      ProcessValue <- "84_Setpoints_PIT402_Main_Target"
   TextField "Text field_27" at 697,736 size 58x20; Text 'Opened'
   TextField "Text field_29" at 306,694 size 300x20; Text 'Air / Inert Gas Pressure Setpoint (Current)'
   AlarmView "Alarm view_1" at 0,777 size 1280x23
   TextField "Text field_6" at 531,373 size 64x18; Text 'Running'
   TextField "Text field_9" at 530,395 size 57x25; Text 'Running'
      Visibility <- "10_DI_Data_E139_RUNNING"
   IOField "I/O field_4" at 917,398 size 89x25; FormatPattern 999999; Unit h
      ProcessValue <- "82_To_HMI_CA Blower Total Run Hours"
   TextField "Text field_30" at 1011,400 size 123x20; Text 'Total Run Hours'
   IOField "I/O field_21" at 916,146 size 90x25; FormatPattern 999999; Unit  h
      ProcessValue <- "82_To_HMI_I&A Compressor Total Run Hours"
   TextField "Text field_31" at 1011,148 size 123x20; Text 'Total Run Hours'
   IOField "I/O field_22" at 935,109 size 40x25; FormatPattern 99; Unit d
      ProcessValue <- "82_To_HMI_P301 CSW Pump Run Days"
   IOField "I/O field_23" at 1068,362 size 40x25; FormatPattern 99; Unit s
      ProcessValue <- "82_To_HMI_CA Blower Run Seconds"

screen "Cooling System" 1280x800, template "Template"
   Group "Group_1" at 335,308 size 88x156; Picture "Graphic_148"
   Group "Group_2" at 298,412 size 194x121; Picture "Graphic_224"
   GraphicView "Graphic view_14" at 335,308 size 85x153; Picture "Graphic_148"
   GraphicView "Graphic view_9" at 298,414 size 189x119; Picture "Graphic_224"
   Group "Group_4" at 1043,404 size 88x156; Picture "Graphic_148"
   Group "Group_5" at 1006,508 size 194x121; Picture "Graphic_224"
   GraphicView "Graphic view_27" at 1043,404 size 85x153; Picture "Graphic_148"
   GraphicView "Graphic view_28" at 1006,511 size 189x119; Picture "Graphic_224"
   Rectangle "Rectangle_7" at 224,48 size 554x250
      Visibility <- "80_From_HMI_P301_PRSNT"
   GraphicView "Graphic view_13" at 501,485 size 115x33; Picture "Graphic_232"
   GraphicView "Graphic view_1" at 446,429 size 75x87; Picture "Graphic_238"
   GraphicView "Graphic view_34" at 489,470 size 52x87; Picture "Graphic_169"
   GraphicView "Graphic view_11" at 80,468 size 424x50; Picture "Graphic_232"
   Group "Group_3" at 298,308 size 194x225; Picture "Graphic_148"
   GraphicView "Graphic view_2" at 480,389 size 43x49; Picture "Graphic_231"
   GraphicView "Graphic view_23" at 832,606 size 29x189; Picture "Graphic_231"
   GraphicView "Graphic view_18" at 802,567 size 88x52; Picture "Graphic_240"
   GraphicView "Graphic view_7" at 175,602 size 43x189; Picture "Graphic_231"
   GraphicView "Graphic view_29" at 964,565 size 56x50; Picture "Graphic_232"
   GraphicView "Graphic view_16" at 1150,564 size 56x50; Picture "Graphic_232"
   GraphicView "Graphic view_10" at 175,547 size 43x16; Picture "Graphic_231"
   GraphicView "Graphic view_8" at 25,514 size 207x209; Picture "Graphic_230"
   Button "HmiScreenItemData_1" at 1,1 size 150x43; TextOn 'Back'; TextOff 'Main Index'
      on Release: ActivateScreen("02 Main Index", 0)
   Rectangle "Rectangle_8" at 237,87 size 528x35
      Visibility <- "80_From_HMI_P301_PRSNT"
   Button "Button_15" at 468,92 size 57x25; TextOn 'Enabled'; TextOff 'Disabled'
      Visibility <- "80_From_HMI_P301_PRSNT"
   Button "Button_16" at 622,92 size 64x25; TextOn 'Alarm'; TextOff 'Text'
      Visibility <- "80_From_HMI_P301_PRSNT"
   TextField "Text field_14" at 239,94 size 185x20; Text 'Cooling Sea Water Pump'
   Button "Button_1" at 545,92 size 57x25; TextOn 'Enabled'; TextOff 'Stopped'
      Visibility <- "80_From_HMI_P301_PRSNT"
   Rectangle "Rectangle_1" at 236,83 size 530x212
      Visibility <- "80_From_HMI_P301_PRSNT"
   TextField "Text field_1" at 387,56 size 235x26; Text 'Cooling System Control'
   TextField "Text field_32" at 468,92 size 57x25; Text 'Enabled'
      Visibility <- "10 DI_DATA_P301_ENBLD"
   TextField "Text field_2" at 543,92 size 59x25; Text 'Running'
      Visibility <- "10_DI_Data_CV311_OPN(1)"
   Button "Button_2" at 622,92 size 64x25; TextOn 'Alarm'; TextOff 'Tripped'
      Visibility <- "10 DI_DATA_P301_TRIPPED"
      Appearance <- "10 DI_DATA_P301_TRIPPED"
   TextField "Text field_72" at 2,524 size 121x38; Text 'Cooling Seawater Inlet'
   GraphicView "Graphic view_17" at 464,297 size 75x99; Picture "Graphic_229"
   GraphicView "Graphic view_4" at 801,333 size 43x255; Picture "Graphic_231"
   GraphicView "Graphic view_5" at 786,305 size 72x46; Picture "Graphic_234"
   GraphicView "Graphic view_6" at 25,472 size 56x43; Picture "Graphic_235"
   TextField "Text field_7" at 12,598 size 58x20; Text 'CV-312'
   TextField "Text field_33" at 352,317 size 54x22; Text 'Closed'
      Visibility <- "10_DI_Data_CV311_CLSD"
   TextField "Text field_3" at 352,317 size 54x22; Text 'Opened'
      Visibility <- "10_DI_Data_CV311_OPN"
   TextField "Text field_71" at 351,343 size 58x20; Text 'CV-311'
   GraphicView "Graphic view_3" at 159,470 size 75x87; Picture "Graphic_239"
   TextField "Text field_5" at 534,295 size 105x38; Text 'To Inert Gas Generator'
   TextField "Text field_69" at 13,624 size 54x22; Text 'Closed'
      Visibility <- "10_DI_Data_CV312_CLSD"
   TextField "Text field_6" at 853,250 size 125x55; Text 'Warm Water From Inert Gas Generator'
   GraphicView "Graphic view_31" at 248,441 size 24x34; Picture "Graphic_36"
   TextField "Text field_17" at 230,422 size 62x20; Text 'PIT-359'
   IOField "I/O field_6" at 226,403 size 68x18; FormatPattern 99.99; Unit  Bar
      ProcessValue <- "12_AI_Data_PIT359_SCALED"
   GraphicView "Graphic view_21" at 849,377 size 88x52; Picture "Graphic_241"
   GraphicView "Graphic view_22" at 848,417 size 43x157; Picture "Graphic_231"
   TextField "Text field_8" at 867,659 size 78x55; Text 'Drain To Oily Bilge Tank'
   GraphicView "Graphic view_25" at 896,422 size 43x134; Picture "Graphic_231"
   GraphicView "Graphic view_26" at 898,526 size 73x87; Picture "Graphic_242"
   Group "Group_6" at 1006,404 size 194x225; Picture "Graphic_148"
   TextField "Text field_12" at 1053,439 size 58x20; Text 'CV-322'
   TextField "Text field_13" at 1054,413 size 54x22; Text 'Closed'
      Visibility <- "10_DI_Data_CV322_CLSD"
   TextField "Text field_19" at 1054,413 size 54x22; Text 'Opened'
      Visibility <- "10_DI_Data_CV322_OPN"
   TextField "Text field_20" at 1190,615 size 88x38; Text 'To Overboard'
   GraphicView "Graphic view_24" at 697,598 size 181x170; Picture "Graphic_230"
   TextField "Text field_9" at 681,704 size 58x20; Text 'CV-321'
   TextField "Text field_11" at 682,678 size 54x22; Text 'Closed'
      Visibility <- "10_DI_Data_CV321_CLSD"
   GraphicView "Graphic view_15" at 244,714 size 40x61; Picture "Graphic_236"
   TextField "Text field_21" at 214,658 size 93x55; Text 'To Existing Flue Gas Scrubber'
   TextField "Text field_70" at 13,624 size 54x22; Text 'Opened'
      Visibility <- "10_DI_Data_CV312_OPN"
   TextField "Text field_10" at 682,678 size 54x22; Text 'Opened'
      Visibility <- "10_DI_Data_CV321_OPN"
   GraphicView "Graphic view_32" at 512,546 size 30x121; Picture "Graphic_147"
   TextField "Text field_4" at 600,529 size 79x55; Text 'Cooling Seawater To GCU'
   GraphicView "Graphic view_19" at 624,477 size 56x43; Picture "Graphic_235"
   GraphicView "Graphic view_33" at 508,659 size 40x61; Picture "Graphic_236"
   TextField "Text field_22" at 481,722 size 79x55; Text 'Cooling Seawater To PGC'
   GraphicView "Graphic view_12" at 891,714 size 40x61; Picture "Graphic_236"
   GraphicView "Graphic view_30" at 1206,568 size 56x43; Picture "Graphic_235"
   GraphicView "Graphic view_35" at 803,244 size 40x61; Picture "Graphic_236"
   Button "HmiScreenItemData_4" at 1129,1 size 150x43; TextOn 'I&A Compressor Ok'; TextOff 'Back'
      on Release: function_efd93a16()
   AlarmView "Alarm view_1" at 0,777 size 1280x23
   Button "HmiScreenItemData_11" at 345,230 size 69x51; TextOn 'RESET'; TextOff 'Reset'; Authorization "Operate"
      on Press: function_b14e0dd5("82_To_HMI_P301 CSW Pump Reset Hours", 0)
   IOField "I/O field_8" at 270,232 size 65x25; FormatPattern 99999; Unit  h
      ProcessValue <- "64_Functioning Hours_P301_IDB_Hours Functioning"
   IOField "I/O field_9" at 270,262 size 65x25; Authorization "Operating Mode"; FormatPattern 99999; Unit  h
      ProcessValue <- "82_To_HMI_P301 CSW Pump Service Time Hours"
   TextField "Text field_23" at 240,231 size 37x20; Text 'Run'
   TextField "Text field_24" at 240,262 size 37x20; Text 'Set'
   TextField "Text field_25" at 283,121 size 141x20; Text 'Service Hour P301'
   Button "HmiScreenItemData_14" at 263,163 size 183x34; TextOn 'Back'; TextOff 'Text'
   IOField "I/O field_17" at 312,167 size 40x25; FormatPattern 99; Unit h
      ProcessValue <- "82_To_HMI_P301 CSW Pump Run Hours"
   IOField "I/O field_18" at 355,167 size 40x25; FormatPattern 99; Unit m
      ProcessValue <- "82_To_HMI_P301 CSW Pump Run Minutes"
   IOField "I/O field_19" at 398,167 size 40x25; FormatPattern 99; Unit s
      ProcessValue <- "82_To_HMI_P301 CSW Pump Run Seconds"
   IOField "I/O field_21" at 245,203 size 90x25; FormatPattern 999999; Unit  h
      ProcessValue <- "82_To_HMI_P301 CSW Pump Total Run Hours"
   TextField "Text field_31" at 340,205 size 123x20; Text 'Total Run Hours'
   Button "Button_17" at 701,92 size 57x25; TextOn 'Alarm'; TextOff 'Service'
      Visibility <- "80_From_HMI_P301_PRSNT"
   Button "Button_9" at 701,92 size 57x25; TextOn 'Alarm'; TextOff 'Service'
      Visibility <- "82_To_HMI_P301 CSW Pump Service Due"
   IOField "I/O field_1" at 270,167 size 40x25; FormatPattern 99; Unit d
      ProcessValue <- "82_To_HMI_P301 CSW Pump Run Days"
   Rectangle "Rectangle_12" at 224,48 size 554x250
      Visibility <- "80_From_HMI_P301_PRSNT"
   Button "HmiScreenItemData_2" at 520,167 size 184x67; TextOn 'FRESH WATER SYSTEM'; TextOff 'Fresh Water System'; Authorization "Operate"
      on Release: ActivateScreen("Fresh Water System", 0)
      Visibility <- "80_From_HMI_P305_PRSNT"
   Button "HmiScreenItemData_3" at 595,392 size 170x41; TextOn 'STOP CSW OVERRUN'; TextOff 'Stop CSW Overrun'; Authorization "Operating Mode"
      on Press: function_b14e0dd5("80_From_HMI_CSW OVR Stop", 0)
      Appearance <- "10_DI_Data_CV311_OPN"

screen "Fresh Water System" 1280x800, template "Template"
   GraphicView "Graphic view_29" at 858,564 size 26x29; Picture "Graphic_155"
   Bar "Bar_1" at 145,436 size 311x274; Unit  %; MinimumValue 0; MaximumValue 100
      ProcessValue <- "12_AI_Data_LIT305_SCALED"
   GraphicView "Graphic view_15" at 640,691 size 216x15; Picture "Graphic_156"
   GraphicView "Graphic view_22" at 468,691 size 71x15; Picture "Graphic_156"
   TextField "Text field_1" at 262,720 size 73x32; Text 'IBC-2 Bulk Tank'
   GraphicView "Graphic view_3" at 454,688 size 6x20; Picture "Graphic_113"
   TextField "Text field_4" at 442,89 size 268x26; Text 'Fresh Water Pump Control'
   IOField "I/O field_2" at 646,242 size 65x25; FormatPattern 99999; Unit  h
      ProcessValue <- "P305_Functioning Hours_IDB_Hours Functioning Out"
   TextField "Text field_5" at 616,244 size 37x20; Text 'Run'
   TextField "Text field_6" at 616,275 size 37x20; Text 'Set'
   TextField "Text field_9" at 659,141 size 100x20; Text 'Service Hour'
   Button "HmiScreenItemData_10" at 639,169 size 178x34; TextOn 'Back'; TextOff 'Text'
   IOField "I/O field_4" at 689,173 size 40x25; FormatPattern 99; Unit h
      ProcessValue <- "82_To_HMI_P305 FW Pump Run Hours"
   IOField "I/O field_5" at 730,173 size 40x25; FormatPattern 99; Unit m
      ProcessValue <- "P305_Functioning Hours_IDB_Minutes"
   IOField "I/O field_6" at 771,173 size 40x25; FormatPattern 99; Unit s
      ProcessValue <- "P305_Functioning Hours_IDB_Seconds"
   Button "Button_4" at 776,90 size 57x25; TextOn 'Alarm'; TextOff 'Service'
      Visibility <- "P305_Functioning Hours_IDB_Service Time bit"
   Button "Button_9" at 374,166 size 57x25; TextOn 'Enabled'; TextOff 'Disabled'
   Button "Button_11" at 528,166 size 64x25; TextOn 'Alarm'; TextOff 'Text'
   TextField "Text field_10" at 231,168 size 140x20; Text 'Fresh Water Pump'
   TextField "Text field_8" at 378,144 size 60x18; Text 'Enabled'
   TextField "Text field_17" at 453,144 size 64x18; Text 'Running'
   TextField "Text field_20" at 533,144 size 58x18; Text 'Tripped'
      Visibility <- "10 DI_DATA_P305_TRIPPED(1)"
   Button "Button_12" at 451,166 size 57x25; TextOn 'Enabled'; TextOff 'Stopped'
   TextField "Text field_26" at 374,166 size 57x25; Text 'Enabled'
      Visibility <- "14_DQ_Data_P305ControlOut"
   TextField "Text field_27" at 448,166 size 64x25; Text 'Running'
      Visibility <- "10 DI_DATA_P305_ENBLD"
   GraphicView "Graphic view_12" at 396,411 size 20x26; Picture "Graphic_36"
   TextField "Text field_11" at 421,411 size 60x18; Text 'LIT-305'
   GraphicView "Graphic view_13" at 518,691 size 71x15; Picture "Graphic_156"
   GraphicView "Graphic view_11" at 456,691 size 15x15; Picture "Graphic_156"
   GraphicView "Graphic view_27" at 846,676 size 25x29; Picture "Graphic_153"
   GraphicView "Graphic view_28" at 858,581 size 13x101; Picture "Graphic_152"
   GraphicView "Graphic view_30" at 876,702 size 146x15; Picture "Graphic_156"
   GraphicView "Graphic view_31" at 870,564 size 152x15; Picture "Graphic_156"
   GraphicView "Graphic view_32" at 858,688 size 26x29; Picture "Graphic_166"
   TextField "Text field_15" at 550,746 size 133x32; Text 'P-305 Fresh Water Pump'
   Button "Button_1" at 528,166 size 64x25; TextOn 'Alarm'; TextOff 'Tripped'
      Visibility <- "10 DI_DATA_P305_TRIPPED"
      Appearance <- "10 DI_DATA_P305_TRIPPED"
   IOField "I/O field_13" at 376,388 size 63x18; FormatPattern 99.9; Unit  %
      ProcessValue <- "12_AI_Data_LIT305_SCALED"
   TextField "Text field_22" at 1059,560 size 168x21; Text 'Fresh Water Supply To GCU'
   TextField "Text field_3" at 1059,699 size 168x21; Text 'Fresh Water Supply To IGG'
   Button "HmiScreenItemData_9" at 721,243 size 69x51; TextOn 'Back'; TextOff 'SReset'; Authorization "Operating Mode"
      on Press: function_b14e0dd5("82_To_HMI_P305 FW Pump Reset Hours", 0)
   GraphicView "Graphic view_1" at 1021,697 size 32x24; Picture "Graphic_244"
   GraphicView "Graphic view_2" at 1021,558 size 32x24; Picture "Graphic_244"
   Button "HmiScreenItemData_1" at 1,1 size 150x43; TextOn 'Back'; TextOff 'Main Index'
      on Release: ActivateScreen("02 Main Index", 0)
   GraphicIOField "Graphic I/O field_3" at 586,670 size 60x65; PictureList "Pump Ani"
      ProcessValue <- "FW Pump Animation"
   Button "HmiScreenItemData_3" at 1129,1 size 150x43; TextOn 'I&A Compressor Ok'; TextOff 'Back'
      on Release: function_efd93a16()
   AlarmView "Alarm view_1" at 0,777 size 1280x23
   IOField "I/O field_21" at 617,211 size 90x25; FormatPattern 999999; Unit  h
      Visibility <- "80_From_HMI_P301_PRSNT"
      ProcessValue <- "P305_Functioning Hours_IDB_Hours Total"
   TextField "Text field_31" at 712,213 size 123x20; Text 'Total Run Hours'
      Visibility <- "80_From_HMI_P301_PRSNT"
   IOField "I/O field_1" at 648,173 size 40x25; FormatPattern 99; Unit d
      ProcessValue <- "82_To_HMI_P305 FW Pump Run Days"
   IOField "I/O field_9" at 646,273 size 65x25; Authorization "Commissioning"; FormatPattern 99999; Unit  h
      Visibility <- "80_From_HMI_P301_PRSNT"
      ProcessValue <- "HMI Data_Fresh Water Service Time"
   Button "HmiScreenItemData_4" at 488,210 size 75x34; TextOn 'STOP'; TextOff 'Stop'
      on Press: ResetBit("80_From_HMI_MAN_DQ_1_7(1)")
   Button "HmiScreenItemData_2" at 385,210 size 75x34; TextOn 'START'; TextOff 'Start'
      on Press: SetBit("80_From_HMI_MAN_DQ_1_7(1)")
   Rectangle "Rectangle_7" at 208,78 size 656x250
      Visibility <- "80_From_HMI_P305_PRSNT"

screen "Fuel System" 1280x800, template "Template"
   GraphicView "Graphic view_4" at 570,430 size 24x23; Picture "Graphic_102"
   Button "HmiScreenItemData_1" at 1,1 size 150x43; TextOn 'Back'; TextOff 'Main Index'
      on Release: ActivateScreen("02 Main Index", 0)
   TextField "Text field_3" at 691,522 size 55x18; Text 'E-500B'
   GraphicView "Graphic view_16" at 658,375 size 123x15; Picture "Graphic_99"
   GraphicIOField "Graphic I/O field_1" at 686,356 size 60x65; PictureList "Pump Ani"
      ProcessValue <- "82_To_HMI_Fuel Pump 1 Animation"
   GraphicView "Graphic view_10" at 657,477 size 124x15; Picture "Graphic_99"
   GraphicIOField "Graphic I/O field_2" at 686,459 size 60x65; PictureList "Pump Ani"
      ProcessValue <- "82_To_HMI_Fuel Pump 2 Animation"
   GraphicView "Graphic view_17" at 642,390 size 15x94; Picture "Graphic_101"
   GraphicView "Graphic view_14" at 643,466 size 21x25; Picture "Graphic_96"
   GraphicView "Graphic view_18" at 643,376 size 24x23; Picture "Graphic_102"
   GraphicView "Graphic view_19" at 638,425 size 18x23; Picture "Graphic_105"
   GraphicView "Graphic view_20" at 782,390 size 15x94; Picture "Graphic_101"
   GraphicView "Graphic view_9" at 772,376 size 24x23; Picture "Graphic_104"
   GraphicView "Graphic view_21" at 771,467 size 25x24; Picture "Graphic_97"
   GraphicView "Graphic view_7" at 783,426 size 19x24; Picture "Graphic_103"
   GraphicView "Graphic view_22" at 578,429 size 71x15; Picture "Graphic_99"
   GraphicView "Graphic view_23" at 789,430 size 94x15; Picture "Graphic_99"
   GraphicView "Graphic view_24" at 672,375 size 18x15; Picture "Graphic_99"
   GraphicView "Graphic view_25" at 672,477 size 18x15; Picture "Graphic_99"
   TextField "Text field_2" at 691,422 size 56x18; Text 'E-500A'
   GraphicView "Graphic view_1" at 621,429 size 27x15; Picture "Graphic_99"
   Button "Button_15" at 157,172 size 57x25; TextOn 'Enabled'; TextOff 'Disabled'
   TextField "Text field_14" at 59,174 size 92x20; Text 'Fuel Pump 1'
   TextField "Text field_15" at 161,151 size 60x18; Text 'Enabled'
   TextField "Text field_18" at 391,149 size 87x18; Text 'Service Due'
   Button "Button_17" at 396,172 size 57x25; TextOn 'Alarm'; TextOff 'Service'
   Button "Button_18" at 159,375 size 57x25; TextOn 'Enabled'; TextOff 'Disabled'
   TextField "Text field_19" at 61,377 size 92x20; Text 'Fuel Pump 2'
   Button "Button_20" at 398,375 size 57x25; TextOn 'Alarm'; TextOff 'Service'
   Rectangle "Rectangle_13" at 678,350 size 77x92
      Appearance <- "10_DI_Data_E500A_TRIPPED"
   Rectangle "Rectangle_14" at 678,453 size 77x92
      Appearance <- "10_DI_Data_E500B_TRIPPED(1)"
   TextField "Text field_7" at 678,544 size 83x18; Text 'Duty Pump'
      Visibility <- "101_Fuel_Pumps_DB_Duty Is B"
   TextField "Text field_12" at 678,333 size 83x18; Text 'Duty Pump'
      Visibility <- "101_Fuel_Pumps_DB_Duty Is A"
   GraphicView "Graphic view_8" at 854,430 size 152x15; Picture "Graphic_99"
   Button "Button_9" at 396,172 size 57x25; TextOn 'Alarm'; TextOff 'Service'
      Visibility <- "82_To_HMI_E500A Fuel Pump Service Due"
   Button "Button_10" at 398,375 size 57x25; TextOn 'Alarm'; TextOff 'Service'
      Visibility <- "82_To_HMI_E500B Fuel Pump Service Due"
   GraphicView "Graphic view_76" at 951,407 size 20x26; Picture "Graphic_36"
   TextField "Text field_23" at 933,442 size 61x18; Text 'PIT-204'
   GraphicView "Graphic view_46" at 997,420 size 20x24; Picture "Graphic_40"
   GraphicView "Graphic view_54" at 1016,372 size 24x21; Picture "Graphic_107"
   TextField "Text field_33" at 1022,392 size 60x18; Text 'TIT-202'
   GraphicView "Graphic view_45" at 1005,315 size 13x117; Picture "Graphic_57"
   TextField "Text field_1" at 1049,301 size 172x18; Text 'IGG Pilot & Main Burner'
   GraphicView "Graphic view_2" at 1006,305 size 20x23; Picture "Graphic_102"
   GraphicView "Graphic view_3" at 549,738 size 6x20; Picture "Graphic_113"
   GraphicView "Graphic view_5" at 557,731 size 25x24; Picture "Graphic_111"
   GraphicView "Graphic view_66" at 568,552 size 15x192; Picture "Graphic_112"
   GraphicView "Graphic view_6" at 568,442 size 15x192; Picture "Graphic_112"
   GraphicView "Graphic view_11" at 551,740 size 15x15; Picture "Graphic_99"
   Button "Button_13" at 157,172 size 57x25; TextOn 'Enabled'; TextOff 'Enabled'
      Visibility <- "10_DI_Data_E500A_ENBLD(1)"
   Button "Button_14" at 159,375 size 57x25; TextOn 'Enabled'; TextOff 'Enabled'
      Visibility <- "10_DI_Data_E500B_ENBLD(1)"
   Button "HmiScreenItemData_7" at 525,369 size 69x51; TextOn 'Back'; TextOff 'PSelect'; Authorization "Operate"
      on Press: function_b14e0dd5("80_From_HMI_SW_DTY_PMP_E500", 0)
   IOField "I/O field_1" at 934,390 size 65x22; FormatPattern 99.99; Unit  Bar
      ProcessValue <- "12_AI_Data_PIT204In_SCALED"
   IOField "I/O field_3" at 312,171 size 65x25; FormatPattern 999999
      ProcessValue <- "64_Functioning Hours_E500A_IDB_Hours Functioning"
   TextField "Text field_5" at 315,149 size 72x18; Text 'Hour Run'
   IOField "I/O field_6" at 314,374 size 65x25; FormatPattern 999999
      ProcessValue <- "64_Functioning Hours_E500B_IDB_Hours Functioning"
   Button "Button_1" at 233,172 size 57x25; TextOn 'Alarm'; TextOff 'Text'
   TextField "Text field_6" at 241,149 size 45x18; Text 'Alarm'
   Button "Button_2" at 235,375 size 57x25; TextOn 'Alarm'; TextOff 'Text'
   Button "Button_3" at 233,172 size 57x25; TextOn 'Alarm'; TextOff 'Tripped'
      Visibility <- "10_DI_Data_E500A_TRIPPED"
      Appearance <- "10_DI_Data_E500A_TRIPPED"
   Button "Button_4" at 235,375 size 57x25; TextOn 'Alarm'; TextOff 'Tripped'
      Visibility <- "10_DI_Data_E500B_TRIPPED(1)"
      Appearance <- "10_DI_Data_E500B_TRIPPED(1)"
   IOField "I/O field_4" at 1043,373 size 55x18; FormatPattern 99.9; Unit  °C
      ProcessValue <- "12_AI_Data_TIT202In_SCALED"
   Button "HmiScreenItemData_3" at 1129,1 size 150x43; TextOn 'I&A Compressor Ok'; TextOff 'Back'
      on Release: function_efd93a16()
   AlarmView "Alarm view_1" at 0,777 size 1280x23
   Button "HmiScreenItemData_11" at 253,294 size 69x51; TextOn 'RESET'; TextOff 'Reset'; Authorization "Operate"
      on Press: function_b14e0dd5("82_To_HMI_E500A Fuel Pump Reset Hours", 0)
   IOField "I/O field_8" at 178,296 size 65x25; FormatPattern 99999; Unit  h
      ProcessValue <- "64_Functioning Hours_E500A_IDB_Hours Functioning"
   IOField "I/O field_9" at 178,326 size 65x25; Authorization "Operate"; FormatPattern 99999; Unit  h
      ProcessValue <- "82_To_HMI_E500A Fuel Pump Service Time Hours"
   TextField "Text field_8" at 148,295 size 37x20; Text 'Run'
   TextField "Text field_21" at 148,326 size 37x20; Text 'Set'
   TextField "Text field_13" at 191,201 size 151x20; Text 'Service Hour E500A'
   Button "HmiScreenItemData_14" at 171,227 size 150x34; TextOn 'Back'; TextOff 'Text'
   IOField "I/O field_17" at 176,231 size 54x25; FormatPattern 999; Unit h
      ProcessValue <- "64_Functioning Hours_E500A_IDB_Hours Functioning"
   IOField "I/O field_18" at 232,231 size 40x25; FormatPattern 99; Unit m
      ProcessValue <- "82_To_HMI_E500A Fuel Pump Run Minutes"
   IOField "I/O field_19" at 275,231 size 40x25; FormatPattern 99; Unit s
      ProcessValue <- "82_To_HMI_E500A Fuel Pump Run Seconds"
   IOField "I/O field_21" at 153,267 size 90x25; FormatPattern 999999; Unit  h
      ProcessValue <- "82_To_HMI_E500A Fuel Pump Total Run Hours"
   TextField "Text field_31" at 248,269 size 123x20; Text 'Total Run Hours'
   Button "HmiScreenItemData_2" at 255,502 size 69x51; TextOn 'RESET'; TextOff 'Reset'; Authorization "Operate"
      on Press: function_b14e0dd5("82_To_HMI_E500B Fuel Pump Reset Hours", 0)
   IOField "I/O field_5" at 180,504 size 65x25; FormatPattern 99999; Unit  h
      ProcessValue <- "64_Functioning Hours_E500B_IDB_Hours Functioning"
   IOField "I/O field_7" at 180,534 size 65x25; Authorization "Operate"; FormatPattern 99999; Unit  h
      ProcessValue <- "82_To_HMI_E500B Fuel Pump Service Time Hours"
   TextField "Text field_9" at 150,503 size 37x20; Text 'Run'
   TextField "Text field_10" at 150,534 size 37x20; Text 'Set'
   TextField "Text field_11" at 193,402 size 149x20; Text 'Service Hour E500B'
   Button "HmiScreenItemData_4" at 174,430 size 150x34; TextOn 'Back'; TextOff 'Text'
   IOField "I/O field_10" at 179,434 size 54x25; FormatPattern 999; Unit h
      ProcessValue <- "64_Functioning Hours_E500B_IDB_Hours Functioning"
   IOField "I/O field_11" at 235,434 size 40x25; FormatPattern 99; Unit m
      ProcessValue <- "82_To_HMI_E500B Fuel Pump Run Minutes"
   IOField "I/O field_12" at 278,434 size 40x25; FormatPattern 99; Unit s
      ProcessValue <- "82_To_HMI_E500B Fuel Pump Run Seconds"
   IOField "I/O field_13" at 155,475 size 90x25; FormatPattern 999999; Unit  h
      ProcessValue <- "82_To_HMI_E500B Fuel Pump Total Run Hours"
   TextField "Text field_16" at 250,477 size 123x20; Text 'Total Run Hours'

screen "IG Transfer Mode" 1280x800, template "Template"
   Group "Group_1" at 596,282 size 37x72; Picture "Graphic_148"
   Group "Group_2" at 581,330 size 80x56; Picture "Graphic_224"
   GraphicView "Graphic view_14" at 596,282 size 36x71; Picture "Graphic_148"
   GraphicView "Graphic view_9" at 581,331 size 78x55; Picture "Graphic_224"
   Group "Group_4" at 670,65 size 37x72; Picture "Graphic_148"
   Group "Group_5" at 655,113 size 80x56; Picture "Graphic_224"
   GraphicView "Graphic view_28" at 670,65 size 36x71; Picture "Graphic_148"
   GraphicView "Graphic view_29" at 655,114 size 78x55; Picture "Graphic_224"
   Group "Group_7" at 302,283 size 37x72; Picture "Graphic_148"
   Group "Group_8" at 287,331 size 80x56; Picture "Graphic_224"
   GraphicView "Graphic view_7" at 302,283 size 36x71; Picture "Graphic_148"
   GraphicView "Graphic view_10" at 287,332 size 78x55; Picture "Graphic_224"
   Group "Group_10" at 871,216 size 37x72; Picture "Graphic_148"
   Group "Group_11" at 856,264 size 80x56; Picture "Graphic_224"
   GraphicView "Graphic view_6" at 871,216 size 36x71; Picture "Graphic_148"
   GraphicView "Graphic view_12" at 856,265 size 78x55; Picture "Graphic_224"
   GraphicView "Graphic view_24" at 761,309 size 18x78; Picture "Graphic_231"
   GraphicView "Graphic view_27" at 472,141 size 336x19; Picture "Graphic_232"
   Group "Group_6" at 655,65 size 80x104; Picture "Graphic_148"
   GraphicView "Graphic view_8" at 454,142 size 31x33; Picture "Graphic_178"
   Group "Group_3" at 581,282 size 80x104; Picture "Graphic_148"
   Button "HmiScreenItemData_1" at 1,1 size 150x43; TextOn 'Back'; TextOff 'Main Index'
      on Release: ActivateScreen("02 Main Index", 0)
   TextField "Text field_5" at 111,336 size 84x55; Text 'From Inert Gas Generator'
   TextField "Text field_12" at 655,72 size 58x20; Text 'CV-432'
   TextField "Text field_13" at 586,268 size 54x22; Text 'Closed'
      Visibility <- "10_DI_Data_CV431_CLSD"
   TextField "Text field_19" at 586,268 size 54x22; Text 'Opened'
      Visibility <- "10_DI_Data_CV431_OPN"
   TextField "Text field_9" at 582,291 size 58x20; Text 'CV-431'
   TextField "Text field_10" at 655,50 size 54x22; Text 'Opened'
      Visibility <- "10_DI_Data_CV432_OPN"
   Button "HmiScreenItemData_17" at 1,46 size 150x43; TextOn 'IGG Plant'; TextOff 'IGGS Plant'
      on Release: ActivateScreen("Inert Gas Generator Plant", 0)
   GraphicView "Graphic view_35" at 696,328 size 264x286; Picture "Graphic_251"
   GraphicView "Graphic view_4" at 749,359 size 30x28; Picture "Graphic_169"
   GraphicView "Graphic view_18" at 759,509 size 25x27; Picture "Graphic_265"
   GraphicView "Graphic view_20" at 759,531 size 35x38; Picture "Graphic_266"
   GraphicView "Graphic view_5" at 992,464 size 168x269; Picture "Graphic_150"
   GraphicView "Graphic view_21" at 773,548 size 216x22; Picture "Graphic_232"
   GraphicView "Graphic view_22" at 976,533 size 20x49; Picture "Graphic_271"
   GraphicView "Graphic view_23" at 1165,476 size 35x22; Picture "Graphic_232"
   GraphicView "Graphic view_25" at 1154,465 size 20x43; Picture "Graphic_271"
   GraphicView "Graphic view_26" at 640,358 size 115x17; Picture "Graphic_232"
   GraphicView "Graphic view_1" at 265,360 size 329x17; Picture "Graphic_232"
   GraphicView "Graphic view_17" at 453,166 size 18x202; Picture "Graphic_231"
   GraphicView "Graphic view_3" at 214,351 size 56x35; Picture "Graphic_279"
   Group "Group_9" at 287,283 size 80x104; Picture "Graphic_148"
   TextField "Text field_49" at 294,291 size 56x18; Text 'CV-401'
   TextField "Text field_50" at 292,268 size 54x22; Text 'Closed'
      Visibility <- "10_DI_Data_CV401_CLSD"
   TextField "Text field_51" at 292,268 size 54x22; Text 'Opened'
      Visibility <- "10_DI_Data_CV401_OPN"
   GraphicView "Graphic view_2" at 791,129 size 20x43; Picture "Graphic_280"
   TextField "Text field_1" at 874,131 size 88x38; Text 'To Cargo Blanketing'
   GraphicView "Graphic view_11" at 816,134 size 56x35; Picture "Graphic_279"
   TextField "Text field_48" at 744,627 size 112x20; Text 'PG Compressor'
      Appearance <- "10_DI_DATA_E_400_NOK"
   TextField "Text field_56" at 1202,508 size 71x18; Text 'For BWTS'
   TextField "Text field_2" at 1068,752 size 38x20; Text 'GCU'
   TextField "Text field_11" at 655,50 size 54x22; Text 'Closed'
      Visibility <- "10_DI_Data_CV432_CLSD"
   Button "HmiScreenItemData_3" at 1129,1 size 150x43; TextOn 'I&A Compressor Ok'; TextOff 'Back'
      on Release: function_efd93a16()
   AlarmView "Alarm view_1" at 0,777 size 1280x23
   GraphicView "Graphic view_83" at 1184,463 size 96x48; Picture "Graphic_235"
   Button "HmiScreenItemData_5" at 1165,453 size 114x70; TextOn 'Back'; TextOff 'Text'
      on Press: ActivateScreen("Balast Water Treatment Plant", 0)
   GraphicView "Graphic view_108" at 6,137 size 95x48; Picture "Left Arow"
   Button "HmiScreenItemData_14" at 5,124 size 106x107; TextOn 'Back'; TextOff 'Text'
      on Press: ActivateScreen("Inert Gas Generator Plant", 0)
   TextField "Text field_21" at 12,193 size 77x34; Text 'Inert Gas Generator'
   GraphicView "Graphic view_13" at 773,292 size 245x19; Picture "Graphic_232"
   GraphicView "Graphic view_15" at 762,293 size 31x33; Picture "Graphic_178"
   GraphicView "Graphic view_16" at 996,280 size 20x43; Picture "Graphic_280"
   TextField "Text field_3" at 1077,283 size 71x38; Text 'Ambient Air Inlet'
   GraphicView "Graphic view_19" at 1021,285 size 56x35; Picture "left small arrow"
   Group "Group_12" at 856,216 size 80x104; Picture "Graphic_148"
   Button "Button_1" at 666,321 size 296x306; TextOff 'Text'
      on Press: ActivateScreen("Inert Gas Conditioning Plant", 0)
   TextField "Text field_4" at 862,225 size 56x18; Text 'CV-441'
   TextField "Text field_6" at 862,202 size 54x22; Text 'Closed'
      Visibility <- "10_DI_DATA_CV441_CLSD"
   TextField "Text field_7" at 862,202 size 54x22; Text 'Opened'
      Visibility <- "10_DI_DATA_CV441_OPN"

screen "O2 Content Monitoring" 1280x800, template "Template"
   TextField "Text field_10" at 20,573 size 128x20; Text 'E600 O2 Content'
   Button "Button_9" at 180,571 size 57x25; TextOn 'Enabled'; TextOff 'Text'
   TextField "Text field_17" at 20,601 size 125x52; Text 'BWT O2 Content Setpoint'
   Button "Button_11" at 180,607 size 57x25; TextOn 'Enabled'; TextOff 'Text'
   TextField "Text field_20" at 153,468 size 171x26; Text 'E600 O2 Content'
   TextField "Text field_12" at 19,646 size 154x20; Text 'Cargo Blanketing O2'
   IOField "I/O field_2" at 177,571 size 74x25; FormatPattern s99.999; Unit %
      ProcessValue <- "12_AI_Data_E600O2ContentIn"
   IOField "I/O field_6" at 180,645 size 66x25; Authorization "Parameter Change"; FormatPattern 99.99; Unit  %
      ProcessValue <- "84_Setpoints_E600_CB_Target"
   TextField "Text field_3" at 484,512 size 160x20; Text 'Burner Fuel Pressure'
   Button "Button_3" at 644,510 size 57x25; TextOn 'Enabled'; TextOff 'Text'
   TextField "Text field_4" at 484,541 size 161x52; Text 'Burner Fuel Pressure Setpoint'
   TextField "Text field_5" at 575,468 size 296x26; Text 'Burner Fuel Control (CV-203)'
   TextField "Text field_6" at 483,585 size 110x20; Text 'Valve Position'
   IOField "I/O field_1" at 642,510 size 71x25; FormatPattern 99.99; Unit  bar
      ProcessValue <- "12_AI_Data_PIT205In_SCALED"
   IOField "I/O field_5" at 642,584 size 71x25; FormatPattern 999.99; Unit  %
      ProcessValue <- "16_AQ_Data_CV203_CNTRL"
   IOField "I/O field_3" at 180,607 size 66x25; Authorization "Parameter Change"; FormatPattern 99.99; Unit %
      ProcessValue <- "84_Setpoints_E600_BWT_Target"
   Button "HmiScreenItemData_3" at 1,1 size 150x43; TextOn 'Back'; TextOff 'Main Index'
      on Release: ActivateScreen("02 Main Index", 0)
   Button "HmiScreenItemData_1" at 1129,1 size 150x43; TextOn 'I&A Compressor Ok'; TextOff 'Back'
      on Release: function_efd93a16()
   AlarmView "Alarm view_1" at 0,777 size 1280x23
   Gauge "Gauge_2" at 258,545 size 210x210; UnitText '%'; CaptionText 'O2 Content'
      Visibility <- "80_From_HMI_CRG_BLNK_MODE"
      ProcessValue <- "12_AI_Data_E600O2ContentIn"
      MaximumValue <- "84_Setpoints_E600_CB_HighHigh"
   TextField "Text field_11" at 975,675 size 257x27; Text 'Proportionate Component PID'
   TextField "Text field_15" at 975,709 size 257x27; Text 'Integrative Component PID'
   TextField "Text field_16" at 975,742 size 257x27; Text 'Derivative Component PID'
   TextField "Text field_19" at 975,553 size 153x27; Text 'Derivation Time'
   TextField "Text field_1" at 977,490 size 153x27; Text 'GAIN'
   TextField "Text field_18" at 975,519 size 153x27; Text 'Integration Time'
   TextField "Text field_2" at 977,588 size 153x27; Text 'Maximum opening'
   Group "Group_16" at 1130,554 size 112x34; Authorization "User administration"; Picture "Graphic_284"; FormatPattern 99
   Switch "Switch_8" at 1223,676 size 32x29; CaptionText 'Switch'; TextOn 'ON'; TextOff 'OFF'; Authorization "User administration"; PictureOff "Design_5_PilotLight_Green_Off"; PictureOn "Design_5_PilotLight_Green_On"
      on Change: InvertBit("84_Setpoints_P_ON")
      ProcessValue <- "84_Setpoints_P_ON"
   Group "Group_15" at 1130,519 size 112x34; Authorization "User administration"; Picture "Graphic_284"; FormatPattern 99
   Switch "Switch_9" at 1223,710 size 32x29; CaptionText 'Switch'; TextOn 'ON'; TextOff 'OFF'; Authorization "User administration"; PictureOff "Design_5_PilotLight_Green_Off"; PictureOn "Design_5_PilotLight_Green_On"
      on Change: InvertBit("84_Setpoints_I_ON")
      ProcessValue <- "84_Setpoints_I_ON"
   Group "Group_3" at 1130,484 size 112x34; Authorization "User administration"; Picture "Graphic_284"; FormatPattern 99
   Switch "Switch_10" at 1223,741 size 32x29; CaptionText 'Switch'; TextOn 'ON'; TextOff 'OFF'; Authorization "User administration"; PictureOff "Design_5_PilotLight_Green_Off"; PictureOn "Design_5_PilotLight_Green_On"
      on Change: InvertBit("84_Setpoints_D_ON")
      ProcessValue <- "84_Setpoints_D_ON"
   Group "Group_1" at 1130,622 size 112x34; Picture "Graphic_284"; Authorization "Commissioning"; FormatPattern 99
   TextField "Text field_21" at 977,622 size 153x27; Text 'Minimum opening'
   Circle "Circle_29" at 30,726 size 20x20
      Appearance <- "Evolving Setpoint_DB_LevelBetter"
   TextField "Text field_22" at 59,722 size 217x27; Text 'O2 content closing Setpoint'
   TrendView "Trend view_1" at 13,53 size 1256x405
      Visibility <- "80_From_HMI_CRG_BLNK_MODE"
      ValueAxis2End <- "84_Setpoints_Max Opening"
      ValueAxis2Begin <- "84_Setpoints_Min Opening"
      ValueAxis1End <- "84_Setpoints_E600_CB_HighHigh"
   TrendView "Trend view_2" at 6,53 size 1267x409
      Visibility <- "80_From_HMI_BWT_BYPASS"
      ValueAxis2End <- "84_Setpoints_Max Opening"
      ValueAxis2Begin <- "84_Setpoints_Min Opening"
      ValueAxis1End <- "84_Setpoints_E600_BWT_HighHigh"
   Gauge "Gauge_3" at 258,545 size 210x210; UnitText '%'; CaptionText 'O2 Content'
      Visibility <- "80_From_HMI_BWT_BYPASS"
      ProcessValue <- "12_AI_Data_E600O2ContentIn"
      MaximumValue <- "84_Setpoints_E600_BWT_HighHigh"
   TextField "Text field_7" at 485,632 size 176x20; Text 'Atomising Air Pressure'
   Button "Button_1" at 650,630 size 57x25; TextOn 'Enabled'; TextOff 'Text'
   TextField "Text field_8" at 485,667 size 180x36; Text 'Pilot Air Press Setpoint'
   Button "Button_2" at 649,666 size 57x25; TextOn 'Enabled'; TextOff 'Text'
   TextField "Text field_9" at 484,742 size 110x20; Text 'Valve Position'
   IOField "I/O field_4" at 642,630 size 71x25; FormatPattern 99.99; Unit  bar
      ProcessValue <- "12_AI_Data_PIT113In_SCALED"
   IOField "I/O field_7" at 642,741 size 71x25; FormatPattern 999.99; Unit  %
      ProcessValue <- "16_AQ_Data_CV111_CNTRL"
   IOField "I/O field_8" at 642,666 size 71x25; Authorization "Commissioning"; FormatPattern 99.99; Unit  bar
      ProcessValue <- "84_Setpoints_PIT113_Pilot_Target"
   Group "Group_2" at 1130,588 size 112x34; Picture "Graphic_284"; Authorization "Commissioning"; FormatPattern 99
   IOField "I/O field_9" at 642,547 size 71x25; Authorization "Commissioning"; FormatPattern 99.99; Unit  bar
      ProcessValue <- "84_Setpoints_PIT205_Target"
   TextField "Text field_13" at 485,704 size 197x36; Text 'Burner Air Press Setpoint'
   Button "Button_4" at 649,703 size 57x25; TextOn 'Enabled'; TextOff 'Text'
   IOField "I/O field_10" at 642,703 size 71x25; Authorization "Commissioning"; FormatPattern 99.99; Unit  bar
      ProcessValue <- "84_Setpoints_PIT113_Burner_Target"
   Gauge "Gauge_4" at 721,547 size 211x211; UnitText '%'; CaptionText 'CV 203'
      ProcessValue <- "16_AQ_Data_CV203_CNTRL"
   GraphicView "Graphic view_22" at 1130,519 size 112x34; Picture "Graphic_284"
   IOField "D5_I/O field_2" at 1145,527 size 62x18; Authorization "User administration"; FormatPattern 99999
      ProcessValue <- "84_Setpoints_Integration Time"
   TextField "D5_Text field_2" at 1205,527 size 23x18; Text 'ms / km/h'
   GraphicView "Graphic view_23" at 1130,554 size 112x34; Picture "Graphic_284"
   IOField "D5_I/O field_3" at 1145,562 size 62x18; Authorization "User administration"; FormatPattern 99999
      ProcessValue <- "84_Setpoints_Derive Time"
   TextField "D5_Text field_3" at 1205,562 size 23x18; Text 'ms / km/h'
   GraphicView "Graphic view_25" at 1130,484 size 112x34; Picture "Graphic_284"
   IOField "D5_I/O field_10" at 1145,492 size 62x18; Authorization "User administration"; FormatPattern 99.9999
      ProcessValue <- "84_Setpoints_Gain"
   TextField "D5_Text field_10" at 1205,492 size 23x18; Text 'km/h'
   GraphicView "Graphic view_1" at 1130,622 size 112x34; Picture "Graphic_284"
   IOField "D5_I/O field_1" at 1145,630 size 62x18; Authorization "Commissioning"; FormatPattern 999; Unit %
      ProcessValue <- "84_Setpoints_Min Opening"
   TextField "D5_Text field_1" at 1205,630 size 23x18; Text 'km/h'
   GraphicView "Graphic view_2" at 1130,588 size 112x34; Picture "Graphic_284"
   IOField "D5_I/O field_5" at 1145,596 size 62x18; Authorization "Commissioning"; FormatPattern 999; Unit %
      ProcessValue <- "84_Setpoints_Max Opening"
   TextField "D5_Text field_5" at 1205,596 size 23x18; Text 'km/h'

screen "41 BWT Ops" 1280x800, template "Template"
   TextField "Text field_74" at 1110,365 size 100x30; Text 'IGGS'
   GraphicIOField "Graphic I/O field_1" at 1110,395 size 100x90; PictureList "IGGS"
      ProcessValue <- "14_DQ_Data_24PF1"
   TextField "Text field_62" at 1120,485 size 80x25; Text 'Disabled'
   TextField "Text field_77" at 1120,485 size 80x25; Text 'Enabled'
      Visibility <- "14_DQ_Data_24PF1"
   Button "Button_8" at 1100,355 size 120x170; TextOff 'Text'
      on Release: ActivateScreen("Inert Gas Generator Plant", 0)
   TextField "Text field_60" at 920,365 size 100x30; Text 'GCU'
   GraphicIOField "Graphic I/O field_4" at 920,395 size 100x90; PictureList "GCU"
      ProcessValue <- "100_GCU_AUTO_SEQ_DB_RNG"
   TextField "Text field_70" at 930,485 size 80x25; Text 'Disabled'
   TextField "Text field_71" at 930,485 size 80x25; Text 'Enabled'
      Visibility <- "100_GCU_AUTO_SEQ_DB_RNG"
   Button "Button_4" at 910,355 size 120x170; TextOff 'Text'
      on Release: ActivateScreen("Inert Gas Conditioning Plant", 0)
   TextField "Text field_65" at 730,365 size 100x30; Text 'PGC'
   TextField "Text field_75" at 740,485 size 80x25; Text 'Disabled'
   TextField "Text field_76" at 740,485 size 80x25; Text 'Enabled'
      Visibility <- "10_DI_DATA_E_400_RUN"
   GraphicView "Graphic view_76" at 730,395 size 100x90; Picture "Graphic_251"
   Button "Button_6" at 720,355 size 120x170; TextOff 'Text'
      on Release: ActivateScreen("PGC System", 0)
   GraphicView "Graphic view_13" at 441,293 size 50x50; Picture "valvevert"
   GraphicView "Graphic view_59" at 199,433 size 518x14; Picture "Graphic_151"
   GraphicView "Logo" at 1,1 size 219x60; Picture "Logo of IGG HMI"
   Button "HmiScreenItemData_1" at 1,50 size 150x43; TextOn 'Back'; TextOff 'Main Index'
      on Release: ActivateScreen("02 Main Index", 0)
   Button "HmiScreenItemData_2" at 1128,64 size 150x43; TextOn 'Back'; TextOff 'BWT Setup'
      on Release: ActivateScreen("Balast Water Treatment Setup", 0)
   DateTimeField "HmiScreenItemData_17" at 1175,0 size 105x30
   DateTimeField "HmiScreenItemData" at 1175,30 size 105x30
   AlarmView "Alarm view_1" at 0,777 size 1280x23
   TextField "Text field_1" at 324,55 size 640x35; Text 'BASIC BARGE TWO TANK CONTROL SYSTEM'
   TextField "Text field_2" at 484,85 size 320x35; Text 'BTCS ENABLED'
      Visibility <- "80_From_HMI_RUN_BTCS"
   TextField "Text field_3" at 484,85 size 320x35; Text 'BTCS DISABLED'
      Visibility <- "80_From_HMI_RUN_BTCS"
   Button "HmiScreenItemData_19" at 700,128 size 570x30; TextOn 'Back'; TextOff 'IGG STEP'; TextList "STEP LIST BTCS"
      ProcessValue <- "2110_BTCS_CNTRL_DB_BTCS_STEP"
   IOField "I/O field_15" at 600,128 size 90x30; Authorization "Commissioning"; FormatPattern 999; Unit  Step
      ProcessValue <- "2110_BTCS_CNTRL_DB_BTCS_STEP"
   Button "HmiScreenItemData_9" at 490,128 size 100x30; TextOn 'Back'; TextOff 'BTCS PLC'
   Button "HmiScreenItemData_3" at 700,168 size 570x30; TextOn 'Back'; TextOff 'IGG STEP'; TextList "STATE LIST BTCS"
      ProcessValue <- "2110_BTCS_CNTRL_DB_BTCS_STATE"
   IOField "I/O field_16" at 600,168 size 90x30; Authorization "Commissioning"; FormatPattern 9; Unit  State
      ProcessValue <- "2110_BTCS_CNTRL_DB_BTCS_STATE"
   Group "Group" at 1100,355 size 120x170; PictureList "IGGS"
   Group "Group_1" at 910,355 size 120x170; PictureList "GCU"
   Group "Group_2" at 720,355 size 120x170; Picture "Graphic_251"
   GraphicView "Graphic view_3" at 506,400 size 50x50; Picture "Graphic_288"
   GraphicView "Graphic view_6" at 346,400 size 50x50; Picture "Graphic_288"
   GraphicView "Graphic view_9" at 615,400 size 50x50; Picture "Graphic_288"
   TextField "Text field_7" at 610,452 size 60x20; Text 'CV-406'
   TextField "Text field_33" at 610,370 size 60x25; Text 'Closed'
      Visibility <- "10_DI_DATA_CV406_CLSD"
   TextField "Text field_14" at 610,370 size 60x25; Text 'Opened'
      Visibility <- "10_DI_DATA_CV406_OPN"
   TextField "Text field_45" at 501,370 size 60x25; Text 'Closed'
      Visibility <- "10_DI_DATA_CV407_CLSD"
   TextField "Text field_11" at 501,370 size 60x25; Text 'Opened'
      Visibility <- "10_DI_DATA_CV407_OPN"
   TextField "Text field_9" at 341,370 size 60x25; Text 'Closed'
      Visibility <- "10_DI_DATA_CV411_CLSD"
   TextField "Text field_10" at 341,370 size 60x25; Text 'Opened'
      Visibility <- "10_DI_DATA_CV411_OPN"
   TextField "Text field_13" at 470,268 size 60x25; Text 'Opened'
      Visibility <- "10_DI_DATA_CV409_OPN"
   TextField "Text field_12" at 470,268 size 60x25; Text 'Closed'
      Visibility <- "10_DI_DATA_CV409_CLSD"
   TextField "Text field_15" at 456,343 size 60x20; Text 'CV-409'
   TextField "Text field_16" at 501,452 size 60x20; Text 'CV-407'
   GraphicView "Graphic view_106" at 444,337 size 14x101; Picture "Graphic_147"
   TextField "Text field_17" at 341,452 size 60x20; Text 'CV-411'
   GraphicView "Graphic view_14" at 444,255 size 14x40; Picture "Graphic_147"
   TextField "Text field_5" at 237,335 size 60x25; Text 'Opened'
      Visibility <- "20_TANKS_IP_DATA_RIO_02_FIRST_TANK_GTT_ISOL_VALVE_OPEN"
   TextField "Text field_6" at 237,335 size 60x25; Text 'Closed'
      Visibility <- "20_TANKS_IP_DATA_RIO_02_FIRST_TANK_GTT_ISOL_VALVE_CLSD"
   TextField "Text field_8" at 238,456 size 60x25; Text 'Opened'
      Visibility <- "20_TANKS_IP_DATA_RIO_02_SECOND_TANK_GTT_ISOL_VALVE_OPEN"
   TextField "Text field_18" at 238,456 size 60x25; Text 'Closed'
      Visibility <- "20_TANKS_IP_DATA_RIO_02_SECOND_TANK_GTT_ISOL_VALVE_CLSD"
   GraphicView "Graphic view_15" at 208,360 size 50x50; Picture "valvevert"
   TextField "Text field_21" at 223,410 size 80x20; Text 'CV-422-2P'
   GraphicView "Graphic view_16" at 211,320 size 14x42; Picture "Graphic_147"
   GraphicView "Graphic view_17" at 209,481 size 50x50; Picture "valvevert"
   TextField "Text field_22" at 224,531 size 80x20; Text 'CV-421-2S'
   GraphicView "Graphic view_18" at 212,405 size 14x79; Picture "Graphic_147"
   GraphicView "Graphic view_11" at 212,527 size 14x33; Picture "Graphic_147"
   Button "Button_1" at 40,130 size 200x150; TextOff 'Tank - 2P'
      Appearance <- "2110_BTCS_CNTRL_DB_PORT_TANK_STS"
   GraphicView "Graphic view_1" at 200,140 size 30x130; Picture "Graphic_183"
   GraphicView "Graphic view_10" at 50,140 size 30x130; Picture "Graphic_183"
   Button "Button_2" at 90,140 size 100x30; TextOff 'Enable / Disable'; TextList "ENBL_DSBL"
      on Press: InvertBit("2110_BTCS_CNTRL_DB_PORT_TANK_STS")
      Appearance <- "2110_BTCS_CNTRL_DB_PORT_TANK_STS"
      ProcessValue <- "2110_BTCS_CNTRL_DB_PORT_TANK_STS"
   Group "Group_3" at 90,240 size 100x20
   Button "Button_7" at 40,600 size 200x150; TextOff 'Tank - 2S'
      Appearance <- "2110_BTCS_CNTRL_DB_STBD_TANK_STS"
   GraphicView "Graphic view_12" at 200,610 size 30x130; Picture "Graphic_183"
   GraphicView "Graphic view_19" at 50,610 size 30x130; Picture "Graphic_183"
   Button "Button_9" at 90,710 size 100x30; TextOff 'Enable / Disable'; TextList "ENBL_DSBL"
      on Press: InvertBit("2110_BTCS_CNTRL_DB_STBD_TANK_STS")
      Appearance <- "2110_BTCS_CNTRL_DB_STBD_TANK_STS"
      ProcessValue <- "2110_BTCS_CNTRL_DB_PORT_TANK_STS"
   Group "Group_4" at 90,615 size 100x20
   TextField "Text field_37" at 5,550 size 90x20; Text 'FIT417 USD'
   IOField "I/O field_10" at 5,570 size 120x25; FormatPattern 9999.9; Unit Nm³/hr
      ProcessValue <- "20_TANKS_IP_DATA_RIO_02_SECOND_TANK_USD_FLOW"
   TextField "Text field_38" at 280,570 size 90x20; Text 'FIT419 MBG'
   IOField "I/O field_11" at 158,570 size 120x25; FormatPattern 9999.9; Unit Nm³/hr
      ProcessValue <- "20_TANKS_IP_DATA_RIO_02_SECOND_TANK_MBG_FLOW"
   TextField "Text field_30" at 5,315 size 90x20; Text 'FIT418 USD'
   IOField "I/O field_5" at 5,290 size 120x25; FormatPattern 9999.9; Unit Nm³/hr
      ProcessValue <- "20_TANKS_IP_DATA_RIO_02_FIRST_TANK_USD_FLOW"
   TextField "Text field_31" at 280,290 size 90x20; Text 'FIT420 MBG'
   IOField "I/O field_6" at 158,290 size 120x25; FormatPattern 9999.9; Unit Nm³/hr
      ProcessValue <- "20_TANKS_IP_DATA_RIO_02_FIRST_TANK_MBG_FLOW"
   IOField "I/O field_30" at 105,355 size 72x25; FormatPattern s999.9; Unit %
      ProcessValue <- "20_TANKS_IP_DATA_RIO_02_FIRST_TANK_BWT_LEVEL"
   IOField "I/O field_31" at 105,483 size 72x25; FormatPattern s999.9; Unit %
      ProcessValue <- "20_TANKS_IP_DATA_RIO_02_SECOND_TANK_BWT_LEVEL"
   IOField "I/O field_32" at 23,355 size 72x25; FormatPattern 999; Unit  DegC
      ProcessValue <- "20_TANKS_IP_DATA_RIO_02_FIRST_TANK_BWT_TEMP"
   IOField "I/O field_33" at 23,483 size 72x25; FormatPattern 999; Unit  DegC
      ProcessValue <- "20_TANKS_IP_DATA_RIO_02_SECOND_TANK_BWT_TEMP"
   IOField "I/O field_34" at 105,386 size 72x25; FormatPattern 9.9; Unit  ph
      ProcessValue <- "20_TANKS_IP_DATA_RIO_02_FIRST_TANK_BWT_PH"
   IOField "I/O field_35" at 105,515 size 72x25; FormatPattern 9.9; Unit  ph
      ProcessValue <- "20_TANKS_IP_DATA_RIO_02_SECOND_TANK_BWT_PH"
   IOField "I/O field_36" at 23,386 size 72x25; FormatPattern 99.9; Unit  mg/l
      ProcessValue <- "20_TANKS_IP_DATA_RIO_02_FIRST_TANK_BWT_DO"
   IOField "I/O field_37" at 23,515 size 72x25; FormatPattern 99.9; Unit  mg/l
      ProcessValue <- "20_TANKS_IP_DATA_RIO_02_SECOND_TANK_BWT_DO"
   IOField "I/O field_2" at 595,481 size 81x25; FormatPattern 999.9; Unit  Barg
      ProcessValue <- "20_TANKS_IP_DATA_RIO_02_FIRST_TANK_DECK_IG_PRESS"
   Button "HmiScreenItemData_4" at 321,635 size 226x75; TextOn 'Back'; TextOff 'MEA Tank Changeover'; TextList "PGC Commissioning"
      on Release: SetBit("PGC_COMMISSION_MODE_DB_Active")
      Visibility <- "10_DI_DATA_E_400_RUN"
      ProcessValue <- "PGC_COMMISSION_MODE_DB_Button Control"
   Circle "Circle_1" at 170,240 size 20x20
      Appearance <- "20_TANKS_IP_DATA_RIO_02_FIRST_TANK_BWT_LEVEL_HIHI"
   TextField "Text field_4" at 90,240 size 75x20; Text 'LS422-2P'
   Circle "Circle_2" at 170,615 size 20x20
      Appearance <- "20_TANKS_IP_DATA_RIO_02_SECOND_TANK_BWT_LEVEL_HIHI"
   TextField "Text field_19" at 90,615 size 75x20; Text 'LS422-2S'

